// TIA Portal project "EdgeHowTos" (V16) (continued)

   // min limit of acutating variable
   IF #statOutput < #minOut THEN
     #statOutput := #minOut;
     #minReached := True;
   ELSE
     #minReached := False;
   END_IF;

   #output := #statOutput;
END_FUNCTION_BLOCK

FUNCTION "Random_Number" : Void   // FC3, SCL
{ S7_Optimized_Access := 'TRUE' }
VERSION : 0.1
   VAR_INPUT
      Min : Int;
      Max : Int;
   END_VAR
   VAR_OUTPUT
      RandomNumber : Int;
   END_VAR
   VAR_TEMP
      range : Int;
      tmp : Int;
   END_VAR
BEGIN
   // generate random number
   #tmp := DINT_TO_INT(TIME_TO_DINT(TIME_TCK()));
   IF #tmp < 0 THEN
       #tmp := #tmp * - 1;
   END_IF;

   "Manipulator" := "Manipulator" + 1;

   IF "Manipulator" = 10 THEN
       "Manipulator" := 1;
   END_IF;

   #tmp := #tmp / "Manipulator";

   #range := #Max - #Min;

   #tmp := #tmp MOD (#range + 1);
   #RandomNumber := #tmp + #Min;
END_FUNCTION

ORGANIZATION_BLOCK "Main"   // OB1, LAD, ProgramCycle
TITLE = "Main Program Sweep (Cycle)"
{ S7_Optimized_Access := 'TRUE' }
VERSION : 0.1
   VAR_INPUT
      Initial_Call : Bool;   // Initial call of this OB
      Remanence : Bool;   // =True, if remanent data are available
   END_VAR
BEGIN
END_ORGANIZATION_BLOCK

ORGANIZATION_BLOCK "Cyclic interrupt"   // OB30, FBD, CyclicInterrupt
{ S7_Optimized_Access := 'TRUE' }
VERSION : 0.1
   VAR_INPUT
      Initial_Call : Bool;   // Initial call of this OB
      Event_Count : Int;   // Events discarded
   END_VAR
BEGIN

REGION Network 1: call filling sequence
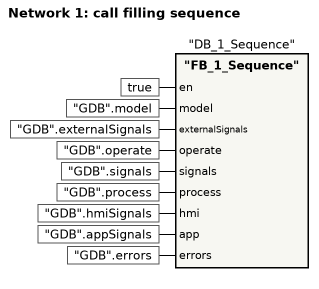
   IF true THEN
       "DB_1_Sequence"(model := "GDB".model,   // "FB_1_Sequence"
                       externalSignals := "GDB".externalSignals,
                       operate := "GDB".operate,
                       signals := "GDB".signals,
                       process := "GDB".process,
                       hmi := "GDB".hmiSignals,
                       app := "GDB".appSignals,
                       errors := "GDB".errors);
   END_IF;
END_REGION
END_ORGANIZATION_BLOCK

(* ===== HMI "HMI_RT_1" =====
system functions are stored by id; their names below are inferred from use

ScreenModuleEditorView "ValueStepperInt_Vertical2" 640x480
   IOField "ioValue" at 0,48 size 80x40; FormatPattern 999999
      ProcessValue <- "value"
   Button "btnIncrease" at 0,0 size 80x40; TextOff 'Text'
      on Click: function_dd21b452("value", "delta")
   Button "btnDecrease" at 0,96 size 80x40; TextOff 'Text'
      on Click: function_b9b71300("value", "delta")
*)

(* ===== HMI "HMI_RT_5" =====
system functions are stored by id; their names below are inferred from use
connection "HMI_Connection_7": 
connection "HMI_Connection_1": ETHERNET, S7_1500_OMS

HMI tags "Template"
   "MainNavigationState" : Int, internal
   "SubNavigationState" : Int, internal
   "CurrentUserName" : WString[18], internal
   "DiagState" : Int, internal
   "PopUpBackground" : Bool, internal
   "UserName" : WString[20], internal
   "Password" : WString[20], internal
   "UserIsLoggedIn" : Bool, internal
   "CodeView" : Bool, internal
   "Brightness" : Int, internal
   "CurrentLanguage" : Bool, internal
   "CurrentRecipeName" : WString[30], internal
   "CurrentMachineState" : Int, internal
   "OptionPanelNavigationState" : Int, internal
   "ButtonDown" : Bool, internal
   "ThirdLevelNavigationState" : Int, internal
   "StartScreenName" : WString[60], internal
   "InScreenTabState" : Int, internal
   "DummyTagBool" : Bool, internal
   "DummyTagInt1" : Int, internal
   "DummyTagInt2" : Int, internal
   "DummyTagInt3" : Int, internal
   "DummyDeltaReal" : LReal, internal
   "DummTagReal1" : LReal, internal
   "DummyDeltaInt" : Int, internal

HMI tags "Filling"
   "hmiStart" : Bool = PLC GDB.hmiSignals.HMI_Start AT %DB1.DBX158.0, 100 ms
   "hmiStop" : Bool = PLC GDB.hmiSignals.HMI_Stop AT %DB1.DBX158.1, 100 ms
   "hmiReset" : Bool = PLC GDB.hmiSignals.HMI_Reset AT %DB1.DBX158.2, 100 ms
   "tankLevel" : Real = PLC GDB.signals.tankSignals.actLevel AT %DB1.DBD94, 100 ms
   "tankTemperature" : Real = PLC GDB.signals.tankSignals.actTemperature AT %DB1.DBD104, 100 ms
   "tankLevelMaxReached" : Bool = PLC GDB.signals.tankSignals.maxLevel AT %DB1.DBX98.0, 100 ms
   "tankTempMax" : Bool = PLC GDB.signals.tankSignals.maxTemperature AT %DB1.DBX108.0, 100 ms
   "hmiNextBottle" : Bool = PLC GDB.hmiSignals.HMI_NextBottle AT %DB1.DBX158.3, 100 ms
   "stateFillingTank" : Bool = PLC GDB.operate.state.FillingTank AT %DB1.DBX2.0, 100 ms
   "stateHeatingTank" : Bool = PLC GDB.operate.state.HeatingTank AT %DB1.DBX2.1, 100 ms
   "stateFillingBottle" : Bool = PLC GDB.operate.state.FillingBottle AT %DB1.DBX2.2, 100 ms
   "stateShiftingBottle" : Bool = PLC GDB.operate.state.ShiftingBottle AT %DB1.DBX2.3, 100 ms
   "stateStop" : Bool = PLC GDB.operate.state.Stop AT %DB1.DBX2.4, 100 ms
   "stateReset" : Bool = PLC GDB.operate.state.Reset AT %DB1.DBX2.5, 100 ms
   "machineState" : Int = PLC GDB.operate.machineState AT %DB1.DBW4, 100 ms
   "tankLevelMax" : Real = PLC GDB.model.tank.maxLevel AT %DB1.DBD22, 100 ms
   "stateRunning" : Bool = PLC DB_1_Sequence.statHmiStateStart, 100 ms
   "bottleID" : UDInt = PLC GDB.process.productId AT %DB1.DBD142, 100 ms
   "bottlesProduced" : UDInt = PLC GDB.process.numberProduced AT %DB1.DBD146, 100 ms
   "bootleNumberFaulty" : UDInt = PLC GDB.process.numberFaulty AT %DB1.DBD150, 100 ms
   "bottleLevel" : Real = PLC GDB.signals.bottleSignals.actLevel AT %DB1.DBD110, 100 ms
   "HMI_bottleLevel1" : Real, internal
   "HMI_bottleLevel2" : Real, internal
   "HMI_bottleLevel3" : Real, internal
   "HMI_bottleLevel" : Real = PLC DB_2_Filling_DB.statHmiBottleLevel AT %DB1.DBD0, 100 ms
   "HMI_doShift" : Bool = PLC DB_2_Filling_DB.statHmiDoShift AT %DB1.DBX0.0, 100 ms
      on ChangeValue: "Conveyor"()
   "qrCode" : String[254] = PLC GDB.appSignals.APP_QRCode AT %DB1.DBX162.0, 100 ms
   "bottleFaulty" : Bool = PLC DB_2_Filling_DB.statHmiFaultyBottle AT %DB1.DBX0.0, 100 ms
   "qrCodeReceived" : Bool = PLC DB_1_Sequence.statHmiQrCodeReceived AT %DB1.DBX0.0, 100 ms
      on ChangeValue: "HandleQrCode"()
   "tempInvisibleObject" : Bool AT %DB1.DBX0.0
   "HMI_bottleInfo1" : Bool AT %DB1.DBX0.0
   "HMI_bottleInfo2" : Bool AT %DB1.DBX0.0
   "HMI_bottleInfo3" : Bool AT %DB1.DBX0.0
   "HMI_bottleInfo4" : Bool AT %DB1.DBX0.0
   "HMI_bottleInfoActive" : Bool, internal
   "energyFillingTank" : Real = PLC GDB.signals.energySignals.energyConsumptionFillingTank AT %DB1.DBD120, 100 ms
   "energyWaterFillingTank" : Real = PLC GDB.signals.energySignals.waterConsumptionFillingTank AT %DB1.DBD124, 100 ms
   "energyHeatingTank" : Real = PLC GDB.signals.energySignals.energyConsumptionHeatingTank AT %DB1.DBD128, 100 ms
   "energyFillingBottles" : Real = PLC GDB.signals.energySignals.energyConsumptionFillingBottles AT %DB1.DBD132, 100 ms
   "tankPressure" : Real = PLC GDB.signals.tankSignals.actPressure AT %DB1.DBD100, 100 ms
   "stateError" : Bool = PLC GDB.operate.state.Error AT %DB1.DBX2.6, 100 ms
   "hmiError" : Bool = PLC GDB.hmiSignals.HMI_Error AT %DB1.DBX158.4, 100 ms
   "alarmIncoming" : Bool = PLC GDB.appSignals.APP_Alarm AT %DB1.DBX418.2, 100 ms
   "batchID" : UDInt = PLC GDB.process.batchId AT %DB1.DBD154, 100 ms
   "energyGas" : Real = PLC GDB.signals.energySignals.gasConsumptionHeatingTank AT %DB1.DBD136, 100 ms

text list "Machine State": 0 'Undefined / Kein Job'; 1 'Production / Produktion'; 2 'Startup / Anlauf'; 3 'Paused / Pausiert'; 4 'Stopped / Gestoppt'; 5 'Shutdown / Beenden'; 6 'Undefined / UNBEKANNT'

text list "timeRange": 1 'Hours / Stunden'; 2 'Days / Tage'; 3 'Weeks / Wochen'; 4 'Months / Monate'; 5 'Years / Jahre'

text list "MachineState_Farfield": 0..1 '???'; 1 'OK'; 2 'ERROR / FEHLER'; 3 'PAUSED / HALT'

text list "Foil Types": 0..1 '120 - 1mm - Transparent'; 1 '120 - 3mm - Transparent'; 2 '240 - 1mm - Transparent'; 3 '240 - 3mm - Transparent'

text list "FunctionState": 0 'Disabled / Deaktiviert'; 1 'Enabled / Aktiviert'

text list "GroundPos": 0 'No / Nein'; 1 'Yes / Ja'

text list "State": 0 'Off / Aus'; 1 'On / An'

graphic list "DiagState": 0 'DiagOkay'; 1 'DiagWarning_1'; 2 'DiagDefault'

graphic list "DiagState_1": 0 'DiagOkay_1'; 1 'DiagWarning'; 2 'DiagDefault'

graphic list "DiagState_2": 0 'DiagOkay_1'; 1 'DiagWarning'; 2 'DiagDefault'

graphic list "DiagState_3": 0 'DiagOkay_White'; 1 'DiagWarning_White'; 2 'Circle'

graphic list "State": 0..1 'OK'; 3 'Error'

graphic list "Machine": 1 'Grafik_Verpackung_Step1_Blink-off'; 2 'Grafik_Verpackung_Step2'; 3 'Grafik_Verpackung_Blink-on'; 6..7 'Grafik_Verpackung_Step1_Blink-off'

screen "30_Diagnostics" 800x480, template "01_One_Nav_Level"
   on GenerateScreen: SetTag("MainNavigationState", 3)
   SysDiagControl "System diagnostics view_1" at 0,104 size 800x375
   GraphicView "Graphic view_2" at 0,0 size 800x480; Picture "PopUpBackground"
      Visibility <- "PopUpBackground"

screen "10_Startscreen" 800x480, template "01_One_Nav_Level"
   on GenerateScreen: "GetStartScreenName"(); SetTag("MainNavigationState", 1)
   GraphicView "Graphic view_2" at 0,0 size 800x480; Picture "PopUpBackground"
      Visibility <- "PopUpBackground"
   GraphicView "bottle finished 1" at 318,346 size 30x70; Picture "Graphic_20"
      Visibility <- "hmiError"
   Bar "Bar_2" at 324,371 size 20x40; MinimumValue 0; MaximumValue 100
      ProcessValue <- "bottleLevel"
      Visibility <- "hmiError"
   GraphicView "bottle finished 1_1" at 279,346 size 30x70; Picture "Graphic_20"
   GraphicView "bottle finished 1_2" at 239,346 size 30x70; Picture "Graphic_20"
   GraphicView "bottle finished 1_3" at 199,346 size 30x70; Picture "Graphic_20"
   Group "Group" at 437,346 size 30x70; Picture "Graphic_20"
   Group "Group_1" at 397,346 size 30x70; Picture "Graphic_20"
   Group "Group_2" at 357,346 size 30x70; Picture "Graphic_20"
   Group "Group_3" at 318,346 size 30x70; Picture "Graphic_20"
   GraphicView "bottle finished 1_4" at 357,346 size 30x70; Picture "Graphic_20"
      Visibility <- "bottlesProduced"
   Bar "Bar_3" at 362,372 size 20x40; MinimumValue 0; MaximumValue 100
      ProcessValue <- "HMI_bottleLevel1"
      Visibility <- "bottlesProduced"
   GraphicView "bottle finished 1_5" at 397,346 size 30x70; Picture "Graphic_20"
      Visibility <- "bottlesProduced"
   Bar "Bar_4" at 402,372 size 20x40; MinimumValue 0; MaximumValue 100
      ProcessValue <- "HMI_bottleLevel2"
      Visibility <- "bottlesProduced"
   GraphicView "bottle finished 1_6" at 437,346 size 30x70; Picture "Graphic_20"
      Visibility <- "bottlesProduced"
   Bar "Bar_5" at 443,372 size 20x40; MinimumValue 0; MaximumValue 100
      ProcessValue <- "HMI_bottleLevel3"
      Visibility <- "bottlesProduced"
   Button "Button_12" at 45,392 size 90x32; TextOn 'Place bottles'; TextOff 'Reset / Place bottle'
      on Press: ResetBit("hmiError")
      Visibility <- "hmiError"
   Rectangle "Rectangle_8" at 682,361 size 88x104
      Visibility <- "HMI_bottleInfoActive"
   GraphicView "Graphic view_4" at 213,87 size 249x237; Picture "Graphic_13"
   Button "Button_4" at 45,159 size 90x48; TextOff 'Start'
      on Press: SetBit("hmiStart")
      on Release: ResetBit("hmiStart")
      Appearance <- "stateRunning"
      ObjectEnable <- "stateRunning"
   Button "Button_5" at 45,215 size 90x48; TextOff 'Stop'
      on Press: SetBit("hmiStop")
      on Release: ResetBit("hmiStop")
      ObjectEnable <- "stateRunning"
      Appearance <- "stateRunning"
   Button "Button_6" at 45,271 size 90x48; TextOff 'Reset'
      on Press: SetBit("hmiReset"); ResetBit("HMI_bottleInfo1"); ResetBit("HMI_bottleInfo2"); ResetBit("HMI_bottleInfo3"); ResetBit("HMI_bottleInfo4"); ResetBit("HMI_bottleInfoActive")
      on Release: ResetBit("hmiReset")
      ObjectEnable <- "stateStop"
      Appearance <- "stateStop"
   IOField "ioKPI" at 700,269 size 68x28; FormatPattern 99.9; Unit  
      ProcessValue <- "tankTemperature"
   IOField "ioKPI_1" at 687,239 size 76x28; FormatPattern 9999
      ProcessValue <- "tankLevel"
   TextField "Text field_3" at 496,160 size 150x25; Text 'Bottles produced'
   Button "Button_1" at 45,354 size 90x32; TextOff 'Reset / Next bottle'
      on Press: SetBit("hmiNextBottle")
      on Release: ResetBit("hmiNextBottle")
      Appearance <- "stateFillingBottle"
      ObjectEnable <- "stateFillingBottle"
   TextField "Text field_1" at 610,106 size 150x25; Text 'Filling tank'
      Visibility <- "stateFillingTank"
   TextField "Text field_5" at 496,106 size 49x25; Text 'State'
   TextField "Text field_6" at 610,106 size 150x25; Text 'Heating tank'
      Visibility <- "stateHeatingTank"
   TextField "Text field_7" at 610,106 size 150x25; Text 'Filling bottle'
      Visibility <- "stateFillingBottle"
   TextField "Text field_8" at 610,106 size 150x25; Text 'Shifting bottle'
      Visibility <- "stateShiftingBottle"
   TextField "Text field_9" at 610,106 size 150x25; Text 'Stop'
      Visibility <- "stateStop"
   TextField "Text field_10" at 610,106 size 150x25; Text 'Reset'
      Visibility <- "stateReset"
   IOField "ioKPI_2" at 638,160 size 124x28; FormatPattern 9999999999
      ProcessValue <- "bottlesProduced"
   TextField "Text field_11" at 496,191 size 119x25; Text 'Bottles faulty'
   IOField "ioKPI_3" at 638,191 size 124x28; FormatPattern 9999999999
      ProcessValue <- "bootleNumberFaulty"
   IOField "ioKPI_4" at 695,329 size 68x28; FormatPattern 999
      ProcessValue <- "bottleLevel"
      Visibility <- "stateShiftingBottle"
   GraphicView "Graphic view_13" at 326,321 size 17x21; Picture "Graphic_18"
   Bar "Bar_1" at 223,115 size 229x206; MinimumValue 0; MaximumValue 1600
      ProcessValue <- "tankLevel"
      Appearance <- "tankTemperature"
   GraphicView "Graphic view_7" at 617,192 size 23x23; Picture "Graphic_58"
      Visibility <- "bottleFaulty"
   IOField "ioKPI_5" at 695,329 size 68x28; FormatPattern 999
      ProcessValue <- "HMI_bottleLevel"
      Visibility <- "stateShiftingBottle"
   Line "Line_1" at 200,422 size 266x0
      Visibility <- "bottlesProduced"
   Rectangle "Rectangle_5" at 356,418 size 32x8
      Visibility <- "bottlesProduced"
   Rectangle "Rectangle_6" at 396,418 size 32x8
      Visibility <- "bottlesProduced"
   Rectangle "Rectangle_7" at 436,418 size 32x8
      Visibility <- "bottlesProduced"
   Line "Line_2" at 200,422 size 225x0
      Visibility <- "bottlesProduced"
   Line "Line_3" at 200,422 size 185x0
      Visibility <- "bottlesProduced"
   Button "Button_2" at 322,431 size 26x22; TextOff 'Text'; PictureOff "Graphic_50"
      on Click: SetBit("HMI_bottleInfo1"); ResetBit("HMI_bottleInfo2"); ResetBit("HMI_bottleInfo3"); ResetBit("HMI_bottleInfo4"); "HandleBottleInfo"()
   Button "Button_7" at 361,431 size 26x22; TextOff 'Text'; PictureOff "Graphic_50"
      on Click: SetBit("HMI_bottleInfo2"); ResetBit("HMI_bottleInfo1"); ResetBit("HMI_bottleInfo3"); ResetBit("HMI_bottleInfo4"); "HandleBottleInfo"()
      Visibility <- "bottlesProduced"
   Button "Button_3" at 400,431 size 26x22; TextOff 'Text'; PictureOff "Graphic_50"
      on Click: SetBit("HMI_bottleInfo3"); ResetBit("HMI_bottleInfo1"); ResetBit("HMI_bottleInfo2"); ResetBit("HMI_bottleInfo4"); "HandleBottleInfo"()
      Visibility <- "bottlesProduced"
   Button "Button_8" at 440,430 size 26x22; TextOff 'Text'; PictureOff "Graphic_50"
      on Click: SetBit("HMI_bottleInfo4"); ResetBit("HMI_bottleInfo1"); ResetBit("HMI_bottleInfo2"); ResetBit("HMI_bottleInfo3"); "HandleBottleInfo"()
      Visibility <- "bottlesProduced"
   IOField "I/O field_1" at 2,459 size 20x20; FormatPattern 1
      Visibility <- "tempInvisibleObject"
      ProcessValue <- "qrCodeReceived"
   GraphicView "Graphic view_1" at 689,384 size 76x76; Picture "QRCode_bottle_one"
      Visibility <- "HMI_bottleInfo1"
   TextField "Text field_2" at 666,359 size 78x25; Text 'bottle 1'
      Visibility <- "HMI_bottleInfo1"
   TextField "Text field_12" at 665,359 size 78x25; Text 'bottle 2'
      Visibility <- "HMI_bottleInfo2"
   GraphicView "Graphic view_3" at 689,384 size 76x76; Picture "QRCode_bottle_two"
      Visibility <- "HMI_bottleInfo2"
   TextField "Text field_13" at 666,359 size 78x25; Text 'bottle 3'
      Visibility <- "HMI_bottleInfo3"
   TextField "Text field_14" at 665,359 size 78x25; Text 'bottle 4'
      Visibility <- "HMI_bottleInfo4"
   GraphicView "Graphic view_5" at 688,384 size 76x76; Picture "QRCode_bottle_three"
      Visibility <- "HMI_bottleInfo3"
   GraphicView "Graphic view_6" at 688,386 size 76x76; Picture "QRCode_bottle_four"
      Visibility <- "HMI_bottleInfo4"
   Button "Button_10" at 501,392 size 100x32; TextOff 'Energy data'; PictureOff "Graphic_50"
      on Click: function_efd93a16("EnergyInfo", 0, 0, -1, -1, 1)
   IOField "ioKPI_6" at 671,299 size 92x28; FormatPattern 999.9
      ProcessValue <- "tankPressure"
   Button "Button_11" at 45,392 size 90x32; TextOn 'Place bottles'; TextOff 'Reset / Push bottle'
      on Press: SetBit("hmiError")
      Visibility <- "hmiError"
   GraphicIOField "D6_Pilotlight_Red" at 92,109 size 40x40; PictureOn "Design_6_PilotLight_Red_On"; PictureOff "Design_6_PilotLight_Red_Off"
      ProcessValue <- "stateError"
   GraphicIOField "D6_Pilotlight_Green" at 48,109 size 40x40; PictureOn "Design_6_PilotLight_Green_On"; PictureOff "Design_6_PilotLight_Green_Off"
      ProcessValue <- "stateRunning"
   TextField "Text field_4" at 610,106 size 150x25; Text 'Error'
      Visibility <- "stateError"
   GraphicView "Graphic view_12" at 138,390 size 28x35; Picture "Graphic_73"
   GraphicView "Graphic view_14" at 138,353 size 28x35; Picture "Graphic_74"
   TextField "Text field_15" at 496,239 size 113x25; Text 'Tank level (l)'
   TextField "Text field_16" at 496,269 size 193x25; Text 'Tank temperature (°C)'
   TextField "Text field_17" at 496,299 size 174x25; Text 'Tank pressure (hPa)'
   TextField "Text field_18" at 496,329 size 124x25; Text 'Bottle level (l)'
   Button "Button_9" at 742,362 size 26x22; TextOff 'Text'; PictureOff "Graphic_68"
      on Click: ResetBit("HMI_bottleInfo1"); ResetBit("HMI_bottleInfo2"); ResetBit("HMI_bottleInfo3"); ResetBit("HMI_bottleInfo4"); ResetBit("HMI_bottleInfoActive")
      Visibility <- "HMI_bottleInfoActive"
   GraphicView "Graphic view_8" at 318,362 size 36x43; Picture "Graphic_72"
      Visibility <- "hmiError"
   Group "Group_4" at 199,346 size 268x70; Picture "Graphic_20"
   IOField "I/O field_2" at 23,459 size 20x20; FormatPattern 1
      Visibility <- "tempInvisibleObject"
      ProcessValue <- "alarmIncoming"
   TextField "Text field_19" at 496,132 size 74x25; Text 'Batch Id'
   IOField "ioKPI_7" at 638,132 size 124x28; FormatPattern 9999999999
      ProcessValue <- "batchID"

Template "01_One_Nav_Level" 800x480
   TextField "txtTitleBar" at 16,8 size 495x32; Text 'Industrial Edge - Tank Application / Applikation'
   Button "btnStartscreen" at 0,0 size 354x45; TextOff 'Text'
      on Click: "ActivateStartScreen"()
   Rectangle "rectSystemDiagnosticsIndicator_1" at 703,0 size 48x48
      Appearance <- "alarmIncoming"
   Rectangle "rectSystemDiagnosticsIndicator" at 752,0 size 48x48
      Appearance <- "DiagState"
   GraphicIOField "gioDiagState" at 760,8 size 32x32; PictureList "DiagState_3"
      ProcessValue <- "DiagState"
   Button "btnDiagState" at 752,0 size 48x48; TextOff 'Text'
      on Click: ActivateScreen("30_Diagnostics", 0)
   TextField "Template_Text field_1" at 720,2 size 17x46; Text '!'
   Button "btnDiagState_1" at 703,0 size 48x48; TextOff 'Text'
      on Click: function_efd93a16("Alarm", 50, 100, -1, -1, 1)

PopupScreen "Template_Logon" 320x352
   on ClearScreen: ResetBit("PopUpBackground")
   on GenerateScreen: SetBit("PopUpBackground")
   TextField "Template_Text field_1" at 16,0 size 215x40; Text 'Login'
   Button "Button_2" at 16,240 size 288x40; TextOn 'LOGIN / ANMELDEN'; TextOff 'LOGIN / ANMELDEN'
      on Click: function_a9b89908("Password", "UserName"); function_efd93a16("Template_Logon", 0, 0, 0, -1, 1)
   IOField "I/O field_1" at 16,84 size 288x40; FormatPattern ??????????????????????????????
      ProcessValue <- "UserName"
   TextField "Text field_1" at 16,56 size 288x24; Text 'User Name / Name'
   IOField "I/O field_2" at 16,168 size 288x40; FormatPattern ??????????????????????????????
      ProcessValue <- "Password"
   TextField "Text field_2" at 16,140 size 288x24; Text 'Password / Passwort'
   Button "Button_1" at 16,296 size 288x40; TextOn 'CLOSE / SCHLIESSEN'; TextOff 'CLOSE / SCHLIESSEN'
      on Click: function_efd93a16("Template_Logon", 0, 0, 0, -1, 1)
      on Press: function_b14e0dd5("ButtonDown", 0)
      Appearance <- "ButtonDown"

PopupScreen "Template_Logon_Logoff" 320x352
   on ClearScreen: ResetBit("PopUpBackground")
   on GenerateScreen: SetBit("PopUpBackground")
   TextField "Template_Text field_1" at 16,0 size 215x40; Text 'Login'
   Button "Button_2" at 16,240 size 136x40; TextOn 'LOG OFF / ABMELDEN'; TextOff 'LOG OFF / ABMELDEN'
      on Click: function_f23ef4c9()
   IOField "I/O field_1" at 16,84 size 288x40; FormatPattern ??????????????????????????????
      ProcessValue <- "UserName"
   TextField "Text field_1" at 16,56 size 288x24; Text 'User Name / Name'
   IOField "I/O field_2" at 16,168 size 288x40; FormatPattern ??????????????????????????????
      ProcessValue <- "Password"
   TextField "Text field_2" at 16,140 size 288x24; Text 'Password / Passwort'
   Button "Button_1" at 16,296 size 288x40; TextOn 'CLOSE / SCHLIESSEN'; TextOff 'CLOSE / SCHLIESSEN'
      on Click: function_efd93a16("Template_Logon_Logoff", 0, 0, 0, -1, 1)
      on Press: function_b14e0dd5("ButtonDown", 0)
      Appearance <- "ButtonDown"
   Button "Button_3" at 168,240 size 136x40; TextOn 'LOGIN / ANMELDEN'; TextOff 'LOGIN / ANMELDEN'
      on Click: function_a9b89908("Password", "UserName"); function_efd93a16("Template_Logon_Logoff", 0, 0, 0, -1, 1)

PopupScreen "Template_Recipe" 700x420
   on ClearScreen: ResetBit("PopUpBackground")
   on GenerateScreen: SetBit("PopUpBackground")
   TextField "Template_Text field_1" at 14,0 size 500x40; Text 'Recipe / Rezeptur'
   Button "Button_1" at 220,364 size 260x40; TextOn 'CLOSE / SCHLIESSEN'; TextOff 'CLOSE / SCHLIESSEN'
      on Click: function_efd93a16("Template_Recipe", 0, 0, 0, -1, 1)
      on Press: function_b14e0dd5("ButtonDown", 0)
      Appearance <- "ButtonDown"
   RecipeView "Rezepturanzeige_1" at 0,40 size 698x320

PopupScreen "OptionPanel_4_Buttons" 400x328
   GraphicView "gfxOptionPanel" at 80,30 size 18x12; Picture "ManFunctions_Off"
   TextField "textOptionPanelTitle" at 108,16 size 260x40; Text 'Option Panel Title / Titel Option Panel'
   Button "btnOptionPanelClose" at 0,0 size 40x328; TextOff 'Text'; PictureOff "Jog_Forward"
      on Press: function_efd93a16("OptionPanel_4_Buttons", 0, 0, 0, 2, 2)
   Button "btnOption1" at 80,72 size 240x40; TextOn 'Option 1'; TextOff 'Option 1 / Move to Home Position'
   Button "btnOption2" at 80,128 size 240x40; TextOn 'Option 2'; TextOff 'Option 2 / Move to Home Position'
   Button "btnOption3" at 80,184 size 240x40; TextOn 'Option 3'; TextOff 'Option 3 / RESET'
   Button "btnOption4" at 80,240 size 240x40; TextOn 'Option 4'; TextOff 'Option 4 / RESET'

SlideinScreen "GraphX_Slidein_Right" 220x480
   Button "Button_1" at 0,78 size 220x60; TextOn 'Menu Item 1'; TextOff 'Startscreen / Startseite'
      on Click: ActivateScreen("10_Startscreen", 0)
      Appearance <- "MainNavigationState"
   Button "Button_3" at 0,201 size 220x60; TextOn 'Menu Item 3'; TextOff 'Diagnostics / Diagnose'
      on Click: ActivateScreen("30_Diagnostics", 0)
      Appearance <- "MainNavigationState"
   Rectangle "Rectangle_1" at 214,78 size 6x60
      Visibility <- "MainNavigationState"
   Rectangle "Rectangle_2" at 214,140 size 6x60
      Visibility <- "MainNavigationState"
   Rectangle "Rectangle_3" at 214,201 size 6x60
      Visibility <- "MainNavigationState"
   Rectangle "Rectangle_4" at 214,262 size 6x60
      Visibility <- "MainNavigationState"

PopupScreen "BottleInfo" 320x352
   on ClearScreen: ResetBit("PopUpBackground")
   on GenerateScreen: SetBit("PopUpBackground")
   TextField "Template_Text field_1" at 16,0 size 215x40; Text 'Bottle information / Login'
   IOField "I/O field_1" at 16,84 size 288x40; FormatPattern 9999
      ProcessValue <- "bottleID"
   TextField "Text field_1" at 16,56 size 288x24; Text 'Production ID / Name'
   IOField "I/O field_2" at 16,168 size 288x40; FormatPattern ??????????????????????????????
      ProcessValue <- "qrCode"
   TextField "Text field_2" at 16,140 size 288x24; Text 'QR Code / Passwort'
   Button "Button_1" at 16,296 size 288x40; TextOn 'CLOSE / SCHLIESSEN'; TextOff 'CLOSE / SCHLIESSEN'
      on Click: function_efd93a16("BottleInfo", 0, 0, 0, -1, 1)
      on Press: function_b14e0dd5("ButtonDown", 0)
      Appearance <- "ButtonDown"

PopupScreen "QRCode" 320x200
   on ClearScreen: ResetBit("PopUpBackground")
   on GenerateScreen: SetBit("PopUpBackground")
   TextField "Template_Text field_1" at 16,0 size 215x40; Text 'QR Code Information / Login'
   IOField "I/O field_2" at 16,64 size 288x40; FormatPattern ??????????????????????????????
      ProcessValue <- "qrCode"
   Button "Button_1" at 16,128 size 288x40; TextOn 'CLOSE / SCHLIESSEN'; TextOff 'CLOSE / SCHLIESSEN'
      on Click: function_efd93a16("QRCode", 0, 0, 0, -1, 1); ResetBit("qrCodeReceived")
      on Press: function_b14e0dd5("ButtonDown", 0)
      Appearance <- "ButtonDown"

PopupScreen "EnergyInfo" 370x352
   on ClearScreen: ResetBit("PopUpBackground")
   on GenerateScreen: SetBit("PopUpBackground")
   IOField "I/O field_3" at 16,248 size 160x40; FormatPattern 9999.99; Unit  Wh
      ProcessValue <- "energyFillingBottles"
   TextField "Template_Text field_1" at 16,0 size 215x40; Text 'Energy consumption / Login'
   IOField "I/O field_1" at 16,103 size 160x40; FormatPattern 9999.99; Unit  Wh
      ProcessValue <- "energyFillingTank"
   TextField "Text field_1" at 16,75 size 152x24; Text 'Filling tank / Name'
   IOField "I/O field_2" at 16,176 size 160x40; FormatPattern 9999.99; Unit  Wh
      ProcessValue <- "energyHeatingTank"
   TextField "Text field_2" at 16,148 size 144x24; Text 'Heating tank / Passwort'
   Button "Button_1" at 16,304 size 344x40; TextOn 'CLOSE / SCHLIESSEN'; TextOff 'CLOSE / SCHLIESSEN'
      on Click: function_efd93a16("EnergyInfo", 0, 0, 0, -1, 1)
      on Press: function_b14e0dd5("ButtonDown", 0)
      Appearance <- "ButtonDown"
   TextField "Text field_3" at 18,220 size 144x24; Text 'Filling bottles / Passwort'
   TextField "Text field_5" at 16,48 size 104x24; Text 'Electricity / Name'
   TextField "Text field_6" at 198,72 size 56x24; Text 'Gas / Name'
   TextField "Text field_4" at 200,147 size 56x24; Text 'Water / Name'
   IOField "I/O field_4" at 200,104 size 160x40; FormatPattern 9999.99; Unit  Wh
      ProcessValue <- "energyGas"
   IOField "I/O field_5" at 200,177 size 160x40; FormatPattern 9999.99; Unit  l
      ProcessValue <- "energyWaterFillingTank"

PopupScreen "Alarm" 700x270
   AlarmView "Alarm view_1" at 5,7 size 688x196
   Button "Button_1" at 192,216 size 288x40; TextOn 'CLOSE / SCHLIESSEN'; TextOff 'CLOSE / SCHLIESSEN'
      on Click: function_efd93a16("Alarm", 0, 0, 0, -1, 1)
      on Press: function_b14e0dd5("ButtonDown", 0)
      Appearance <- "ButtonDown"

VB script "ActivateStartScreen"
   HmiRuntime.BaseScreenName = SmartTags("StartScreenName")

VB script "CheckDiagState"
   If SmartTags("@DiagnosticsIndicatorTag") = 1 Then
   	SmartTags("DiagState") = 1
   Else
   	SmartTags("DiagState") = 0
   End If

VB script "GetStartScreenName"
   SmartTags("StartScreenName") = HmiRuntime.BaseScreenName

VB script "Conveyor"
   ' ---------------- conveyor with bottles ---------------------------
   
   Dim HMI_doShift
   Set HMI_doShift = HmiRuntime.SmartTags("HMI_doShift")
   
   If HMI_doShift.Value = True Then	
   	
   	'Timer - wait to get current value from runtime
   '	Dim counter
   '	counter = 0
   '	While counter < 500
   '		counter = counter +1
   '	Wend
   
   	Dim HMI_bottleLevel
   	Dim HMI_bottleLevel1
   	Dim HMI_bottleLevel3
   	Dim HMI_bottleLevel2
   	
   	Set HMI_bottleLevel = HmiRuntime.SmartTags("HMI_bottleLevel")
   	Set HMI_bottleLevel1 = SmartTags("HMI_bottleLevel1")
   	Set HMI_bottleLevel2 = SmartTags("HMI_bottleLevel2")
   	Set HMI_bottleLevel3 = SmartTags("HMI_bottleLevel3")
   	
   	HMI_bottleLevel3.Value = HMI_bottleLevel2.Value
   	HMI_bottleLevel2.Value = HMI_bottleLevel1.Value	
   	HMI_bottleLevel1.Value = HMI_bottleLevel.Value
   
   End If

VB script "HandleQrCode"
   Dim qrCodeReceived
   Set qrCodeReceived = HmiRuntime.SmartTags("qrCodeReceived")
   
   If qrCodeReceived.Value = True Then	
   	efd93a16-2665-4b85-bcb9-25eddcb7b6f4 QRCode,0,0,$3$hmiOn$,$3$hmiAnimationOff$,$3$hmiFast$
   End If

VB script "TEMPLATE_HandleControls"
   ' ---------------- button "Next bottle" ---------------------------
   ' => if stateFillingBottle
   
   'read value from tag
   'Dim stateFillingBottle
   'Dim buttonNextBottle
   
   'Set stateFillingBottle = HmiRuntime.SmartTags("stateFillingBottle")
   'Set buttonNextBottle = SmartTags("activateButtonNextBottle")
   
   'If stateStop.Value = True And maxTemp.Value = True Then
   'If stateFillingBottle.Value = True Then
   '	buttonNextBottle.Value = True
   'Else
   '	buttonNextBottle.Value = False
   'End If

VB script "HandleBottleInfo"
   Dim HMI_bottleInfo1
   Dim HMI_bottleInfo2
   Dim HMI_bottleInfo3
   Dim HMI_bottleInfo4
   Dim HMI_bottleInfoActive
   
   Set HMI_bottleInfo1 = SmartTags("HMI_bottleInfo1")
   Set HMI_bottleInfo2 = SmartTags("HMI_bottleInfo2")
   Set HMI_bottleInfo3 = SmartTags("HMI_bottleInfo3")
   Set HMI_bottleInfo4 = SmartTags("HMI_bottleInfo4")
   Set HMI_bottleInfoActive = SmartTags("HMI_bottleInfoActive")
   
   
   If (HMI_bottleInfo1.Value = True) Or (HMI_bottleInfo2.Value = True) Or (HMI_bottleInfo3.Value = True) Or (HMI_bottleInfo4.Value = True)  Then	
   	HMI_bottleInfoActive.Value = True
   Else
   	HMI_bottleInfoActive.Value = False
   End If
*)